           // ===============================================================
           // (7) SCAN REFERENCE ACQUISITION — pág. 10
           // FÍSICO: KUKA carga PN/frame y se coloca en el punto de INICIO de
           // la trayectoria de referencia. Tu lógica pone AtRefScanStart=TRUE cuando
           // está en posición. El PLC solo arma scan_ref_start si además los
           // parámetros mínimos (id_scan, x_size, y_size) están válidos (p. 10).
           // ===============================================================
       #cSTEP_SCAN_REF:

           // Validación mínima de parámetros de scan que el PLC publica al Supervisor
           #validScanParams := (LEN("PlcStatus".idScan) > 0) AND ("PlcStatus".xSize > 0.0) AND ("PlcStatus".ySize > 0.0);

           // Posicionar al inicio de Ref si no estamos (CASE 420, ARG=RefProgIdx)
           IF (NOT #kukaAtRefScanStartPos) AND (#WantCode_uint = 0) THEN
               #SupervisorCmdSeq := #SupervisorCmdSeq + 1;
               #WantCode_uint := #cKUKA_GOTO_REF_START; // ← KRC: CASE 420
               #WantProgRequestId := (#RefProgIdx);   // índice de programa REF por pieza
           END_IF;

           // Permiso de arranque
           IF #kukaAtRefScanStartPos AND #validScanParams AND NOT "SupervisorCmd".scanRefRunning THEN
               "PlcStatus".scanRefStart := TRUE;   // ← Anunciar “ready” al Supervisor
           END_IF;

           // Cuando el Supervisor arranca por primera vez → ejecutar trayectoria (CASE 432)
           IF (NOT #scanRefWasRunning) AND "SupervisorCmd".scanRefRunning THEN
               #SupervisorCmdSeq := #SupervisorCmdSeq + 1;
               #WantCode_uint := #cKUKA_RUN_REF_PATH;
               #WantProgRequestId := (#RefProgIdx);
           END_IF;

           IF "SupervisorCmd".scanRefRunning THEN
               #scanRefWasRunning := TRUE;
               IF #kukaRefScanFinished THEN
                   "PlcStatus".scanRefStart := FALSE;
               END_IF;
           END_IF;

           IF (NOT "SupervisorCmd".scanRefRunning) AND #scanRefWasRunning THEN
               #scanRefWasRunning := FALSE;
               "PlcStatus".scanRefStart := FALSE;

               IF NOT "SupervisorCmd".scanRefState THEN
                   "PlcStatus".stepPlc := #cSTEP_ID;
               ELSE
                   "PlcStatus".stepPlc := #cSTEP_SCAN_INSP;
               END_IF;
           END_IF;

           // ===============================================================
           // (8) SCAN INSPECTION — pág. 11
           // FÍSICO: KUKA se coloca en INICIO de la(s) trayectoria(s) de inspección
           // (AtInspScanStart=TRUE). El PLC arma scan_insp_start solo si parámetros
           // válidos. Supervisor corre/guarda y luego pide verificación (req_verif) (p. 11).
           // ===============================================================
       #cSTEP_SCAN_INSP:

           #validScanParams := (LEN("PlcStatus".idScan) > 0) AND ("PlcStatus".xSize > 0.0) AND ("PlcStatus".ySize > 0.0);

           // Posicionar al inicio de Insp (CASE 421, ARG=PartProgIdx)
           IF (NOT #kukaAtInspScanStartPos) AND (#WantCode_uint = 0) THEN
               #SupervisorCmdSeq := #SupervisorCmdSeq + 1;
               #WantCode_uint := #cKUKA_GOTO_INSP_START;
               #WantProgRequestId := (#PartProgIdx);
           END_IF;

           // Permiso de arranque
           IF #kukaAtInspScanStartPos AND #validScanParams AND NOT "SupervisorCmd".scanInsprunning THEN
               "PlcStatus".scanInspStart := TRUE;
           END_IF;

           // Al arrancar por primera vez → ejecutar trayectoria (CASE 433)
           IF (NOT #scanInspWasRunning) AND "SupervisorCmd".scanInsprunning THEN
               #SupervisorCmdSeq := #SupervisorCmdSeq + 1;
               #WantCode_uint := #cKUKA_RUN_INSP_PATH;
               #WantProgRequestId := (#PartProgIdx);
           END_IF;

           IF "SupervisorCmd".scanInsprunning THEN
               #scanInspWasRunning := TRUE;
               IF #kukaInspScanFinished THEN
                   "PlcStatus".scanInspStart := FALSE;
               END_IF;
           END_IF;

           IF (NOT "SupervisorCmd".scanInsprunning) AND #scanInspWasRunning THEN
               #scanInspWasRunning := FALSE;
               "PlcStatus".scanInspStart := FALSE;

               IF NOT "SupervisorCmd".scanInspState THEN
                   "PlcStatus".stepPlc := #cSTEP_ID;
               ELSE
                   // Pasar a verificación (latch)
                   IF "SupervisorCmd".reqVerif AND NOT #L_reqVerif THEN
                       "PlcStatus".stepPlc := #cSTEP_SCAN_REF_VERIF;
                       #L_reqVerif := TRUE;
                   END_IF;
                   IF NOT "SupervisorCmd".reqVerif THEN
                       #L_reqVerif := FALSE;
                   END_IF;
               END_IF;
           END_IF;


           // ===============================================================
           // (9) SCAN REFERENCE VERIFICATION — pág. 12
           // FÍSICO: KUKA vuelve al INICIO de la trayectoria de verificación de ref.
           // (AtRefScanStart=TRUE). Igual patrón de parámetros/ready/running/state (p. 12).
           // Fin: Supervisor decide Pre‑eval (req_pre_eval) o nuevo ciclo (req_identification_state).
           // ===============================================================
       #cSTEP_SCAN_REF_VERIF:

           #validScanParams := (LEN("PlcStatus".idScan) > 0) AND ("PlcStatus".xSize > 0.0) AND ("PlcStatus".ySize > 0.0);

           // Asegurar estar en inicio de Ref (CASE 420) antes de verificar
           IF (NOT #kukaAtRefScanStartPos) AND (#WantCode_uint = 0) THEN
               #SupervisorCmdSeq := #SupervisorCmdSeq + 1;
               #WantCode_uint := #cKUKA_GOTO_REF_START;
               #WantProgRequestId := (#RefProgIdx);
           END_IF;

           IF #kukaAtRefScanStartPos AND #validScanParams AND NOT "SupervisorCmd".scanRefRunning THEN
               "PlcStatus".scanRefStart := TRUE;
           END_IF;

           IF "SupervisorCmd".scanRefRunning THEN
               #scanRefWasRunning := TRUE;
           END_IF;

           IF (NOT "SupervisorCmd".scanRefRunning) AND #scanRefWasRunning THEN
               #scanRefWasRunning := FALSE;
               "PlcStatus".scanRefStart := FALSE;

               IF NOT "SupervisorCmd".scanRefState THEN
                   "PlcStatus".stepPlc := #cSTEP_ID;
               ELSE
                   // a) Pre‑eval
                   IF "SupervisorCmd".reqPreEval AND NOT #L_reqPreEval THEN
                       "PlcStatus".stepPlc := #cSTEP_PRE_EVAL;
                       #L_reqPreEval := TRUE;
                   END_IF;
                   IF NOT "SupervisorCmd".reqPreEval THEN
                       #L_reqPreEval := FALSE;
                   END_IF;

                   // b) Nuevo ciclo
                   IF "SupervisorCmd".reqIdentificationState AND NOT #L_reqIdent THEN
                       "PlcStatus".stepPlc := #cSTEP_ID;
                       #L_reqIdent := TRUE;
                   END_IF;
                   IF NOT "SupervisorCmd".reqIdentificationState THEN
                       #L_reqIdent := FALSE;
                   END_IF;
               END_IF;
           END_IF;

           // ===============================================================
           // (10) PRE‑EVALUATION / MARKING — pág. 13
           // FÍSICO: si la herramienta de marcado no está montada, el KUKA cambia
           // en Staübli al stand de “marking” según requiera el proceso; tras estar
           // listo se puede marcar (Supervisor.req_mark). El resultado físico del
           // marcado tu lógica lo refleja en MarkingDone=TRUE/FALSE (p. 13).
           // También se puede arrancar un nuevo ciclo (req_identification_state).
           // ===============================================================
       #cSTEP_PRE_EVAL:

           // Volver a Identification (una sola vez)
           IF "SupervisorCmd".reqIdentificationState AND NOT #L_reqIdent THEN
               "PlcStatus".stepPlc := #cSTEP_ID;
               #L_reqIdent := TRUE;
           END_IF;
           IF NOT "SupervisorCmd".reqIdentificationState THEN
               #L_reqIdent := FALSE;
           END_IF;

           // Marcado: un ciclo de ejecución por petición
           IF "SupervisorCmd".reqMark AND NOT #L_reqMark THEN
               "PlcStatus".markState := FALSE;
               "PlcStatus".markRunning := TRUE;
               "PlcStatus".markState := #MarkingDone;   // resultado físico del efector
               "PlcStatus".markRunning := FALSE;
               #L_reqMark := TRUE;
           END_IF;
           IF NOT "SupervisorCmd".reqMark THEN
               #L_reqMark := FALSE;
           END_IF;
       ELSE
           "PlcStatus".stepPlc := #cSTEP_ID;


   END_CASE;


   // ---------------------------------------------------------------
   // [2] DESPACHO AL KUKA (toggle goTrigger cuando el canal esté libre)
   //     • Este bloque “consume” el slot WantCmd → publica parámetros
   //       en los registros PNIO (con SWAP) → toggle de goTrigger.
   //     • El robot deberá igualar rbDone := goTrigger al terminar.
   // ---------------------------------------------------------------

   CASE #state OF
       0: // IDLE -> GO == ACK

           // "cancelGo" := FALSE;

           IF (#SupervisorCmdSeq <> #lastSeq) THEN

               IF  "goTrigger" = "rbDone" THEN

                   #code_int := #WantCode_uint;  // “code_int” que viajará al KRC

                   IF #code_int = 201 THEN
                       // id de herramienta → WORD+SWAP
                       // #Cfg_EndEffector
                       #toolReqId := SWAP(INT_TO_WORD(#WantToolRequestId));

                   END_IF;

                   IF #code_int = 414 THEN  //GOTO_TCG
                       // id de herramienta → WORD+SWAP
                       "requestIndexKuka" := SWAP(UINT_TO_WORD(#WantIndex));

                   END_IF;

                   IF #code_int = 420 THEN // GOTO_REF_START
                       // id de herramienta → WORD+SWAP
                       "programReqId" := SWAP(UINT_TO_WORD(#WantProgRequestId));

                   END_IF;

                   IF #code_int = 432 THEN // RUN_REF_PATH
                       // id de herramienta → WORD+SWAP
                       "programReqId" := SWAP(UINT_TO_WORD(#WantProgRequestId));

                   END_IF;

                   IF #code_int = 421 THEN // GOTO_REF_START
                       // id de herramienta → WORD+SWAP
                       "programReqId" := SWAP(UINT_TO_WORD(#WantProgRequestId));

                   END_IF;

                   IF #code_int = 433 THEN // RUN_INSP_PATH

                       "programReqId" := SWAP(UINT_TO_WORD(#WantProgRequestId));

                   END_IF;

                   // 2) Publicar código de movimiento
                   #moveCodeKuka := SWAP(UINT_TO_WORD(#code_int));   // KRC leerá "MoveCode" = INT

                   // 3) Disparo del GO: toggle de goTrigger (rbDone ≠ goTrigger → pedido activo)
                   "goTrigger" := NOT "goTrigger";

                   #lastSeq := #SupervisorCmdSeq;          // <-- memoriza!
                   #state := 20;

               END_IF;
           END_IF;

       20: // BUSY

           //#code_int := #KukaControlCmdCode;

           // CANCEL pedido en BUSY → avisar al KRC y ACK de la ORDEN ACTIVA
           IF #code_int = 903 THEN
               "cancelGo" := TRUE;
           END_IF;

           // Fin normal (o tras el cancel, cuando KRC cierra el canal por nivel)

           IF ("rbDone" = "goTrigger") THEN
               // 4) Vaciar slot de pendiente
               #WantCode_uint := 0;
               #WantProgRequestId := 0;
               #WantToolRequestId := 0;
               #WantIndex := 0;
               #state := 0;                            // vuelve a IDLE
           END_IF;

   END_CASE;
END_REGION
END_FUNCTION_BLOCK

ORGANIZATION_BLOCK "Main"   // OB1, LAD, ProgramCycle
TITLE = "Main Program Sweep (Cycle)"
{ S7_Optimized_Access := 'TRUE' }
VERSION : 0.1
   VAR_INPUT
      Initial_Call : Bool;   // Initial call of this OB
      Remanence : Bool;   // =True, if remanent data are available
   END_VAR
   VAR_TEMP
      evtEnterSrv : Bool;   // // Eventos de modo service jog
      evtEnterAuto : Bool;   // // Eventos de modo auto
      muxSelStb : Bool;
      muxStartStb : Bool;
      muxPgno : Byte;
      u : UDInt;
   END_VAR
BEGIN

REGION Network 1 (SCL): // ====================== READ (%I) ======================
   // // —— Enlaza estos símbolos a tus %I en el árbol de dispositivos ——
   //   // EStop_DI, SafeDoor_DI, AirPressure_DI, WaterInsp_DI, WaterTank_DI, RobotReady_DI, ...
   "$MOVE_ENABLE" := TRUE;
   "$I_O_ACT" := TRUE;
   //"$IN_HOME"
   //"$EXT"
   "PlcStatus".systemArmed := FALSE;
   "PlcStatus".robotInAutExt := "$EXT";
   "PlcStatus".robotInHome := "$IN_HOME";
END_REGION

REGION Network 2
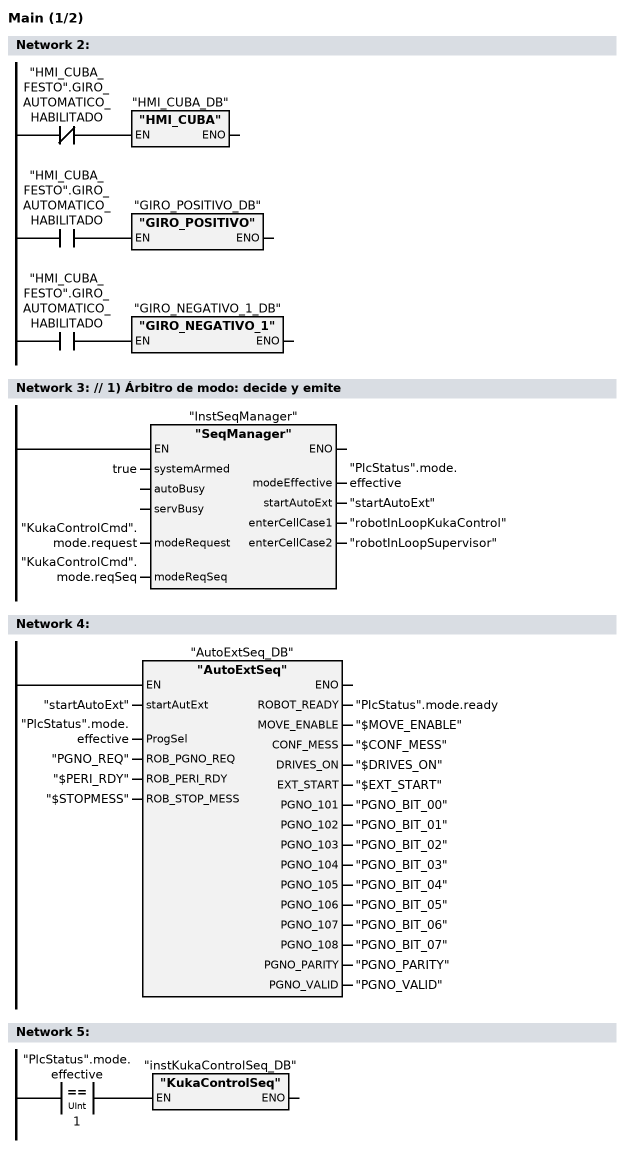
   RUNG wire#powerrail
      I_Contact( "HMI_CUBA_FESTO".GIRO_AUTOMATICO_HABILITADO )
      "HMI_CUBA_DB"()
   END_RUNG
   RUNG wire#powerrail
      Contact( "HMI_CUBA_FESTO".GIRO_AUTOMATICO_HABILITADO )
      "GIRO_POSITIVO_DB"()
   END_RUNG
   RUNG wire#powerrail
      Contact( "HMI_CUBA_FESTO".GIRO_AUTOMATICO_HABILITADO )
      "GIRO_NEGATIVO_1_DB"()
   END_RUNG
   // the same network as SCL:
   IF NOT "HMI_CUBA_FESTO".GIRO_AUTOMATICO_HABILITADO THEN
       "HMI_CUBA_DB"();   // "HMI_CUBA"
   END_IF;
   IF "HMI_CUBA_FESTO".GIRO_AUTOMATICO_HABILITADO THEN
       "GIRO_POSITIVO_DB"();   // "GIRO_POSITIVO"
   END_IF;
   IF "HMI_CUBA_FESTO".GIRO_AUTOMATICO_HABILITADO THEN
       "GIRO_NEGATIVO_1_DB"();   // "GIRO_NEGATIVO_1"
   END_IF;
END_REGION

REGION Network 3: // 1) Árbitro de modo: decide y emite
   RUNG wire#powerrail
      "InstSeqManager"(systemArmed := true, autoBusy :=, servBusy :=, modeRequest := "KukaControlCmd".mode.request, modeReqSeq := "KukaControlCmd".mode.reqSeq, modeEffective => "PlcStatus".mode.effective, startAutoExt => "startAutoExt", enterCellCase1 => "robotInLoopKukaControl", enterCellCase2 => "robotInLoopSupervisor")
   END_RUNG
   // the same network as SCL:
   "InstSeqManager"(systemArmed := true,   // "SeqManager"
                    modeRequest := "KukaControlCmd".mode.request,
                    modeReqSeq := "KukaControlCmd".mode.reqSeq,
                    modeEffective => "PlcStatus".mode.effective,
                    startAutoExt => "startAutoExt",
                    enterCellCase1 => "robotInLoopKukaControl",
                    enterCellCase2 => "robotInLoopSupervisor");
END_REGION

REGION Network 4
   RUNG wire#powerrail
      "AutoExtSeq_DB"(startAutExt := "startAutoExt", ProgSel := "PlcStatus".mode.effective, ROB_PGNO_REQ := "PGNO_REQ", ROB_PERI_RDY := "$PERI_RDY", ROB_STOP_MESS := "$STOPMESS", ROBOT_READY => "PlcStatus".mode.ready, MOVE_ENABLE => "$MOVE_ENABLE", CONF_MESS => "$CONF_MESS", DRIVES_ON => "$DRIVES_ON", EXT_START => "$EXT_START", PGNO_101 => "PGNO_BIT_00", PGNO_102 => "PGNO_BIT_01", PGNO_103 => "PGNO_BIT_02", PGNO_104 => "PGNO_BIT_03", PGNO_105 => "PGNO_BIT_04", PGNO_106 => "PGNO_BIT_05", PGNO_107 => "PGNO_BIT_06", PGNO_108 => "PGNO_BIT_07", PGNO_PARITY => "PGNO_PARITY", PGNO_VALID => "PGNO_VALID")
   END_RUNG
   // the same network as SCL:
   "AutoExtSeq_DB"(startAutExt := "startAutoExt",   // "AutoExtSeq"
                   ProgSel := "PlcStatus".mode.effective,
                   ROB_PGNO_REQ := "PGNO_REQ",
                   ROB_PERI_RDY := "$PERI_RDY",
                   ROB_STOP_MESS := "$STOPMESS",
                   ROBOT_READY => "PlcStatus".mode.ready,
                   MOVE_ENABLE => "$MOVE_ENABLE",
                   CONF_MESS => "$CONF_MESS",
                   DRIVES_ON => "$DRIVES_ON",
                   EXT_START => "$EXT_START",
                   PGNO_101 => "PGNO_BIT_00",
                   PGNO_102 => "PGNO_BIT_01",
                   PGNO_103 => "PGNO_BIT_02",
                   PGNO_104 => "PGNO_BIT_03",
                   PGNO_105 => "PGNO_BIT_04",
                   PGNO_106 => "PGNO_BIT_05",
                   PGNO_107 => "PGNO_BIT_06",
                   PGNO_108 => "PGNO_BIT_07",
                   PGNO_PARITY => "PGNO_PARITY",
                   PGNO_VALID => "PGNO_VALID");
END_REGION

REGION Network 5
   RUNG wire#powerrail
      { S7_Templates := "SrcType := UInt" } EQ_Contact(in1 := "PlcStatus".mode.effective, in2 := 1)
      "instKukaControlSeq_DB"()
   END_RUNG
   // the same network as SCL:
   IF "PlcStatus".mode.effective = 1 THEN
       "instKukaControlSeq_DB"();   // "KukaControlSeq"
   END_IF;
END_REGION

REGION Network 6
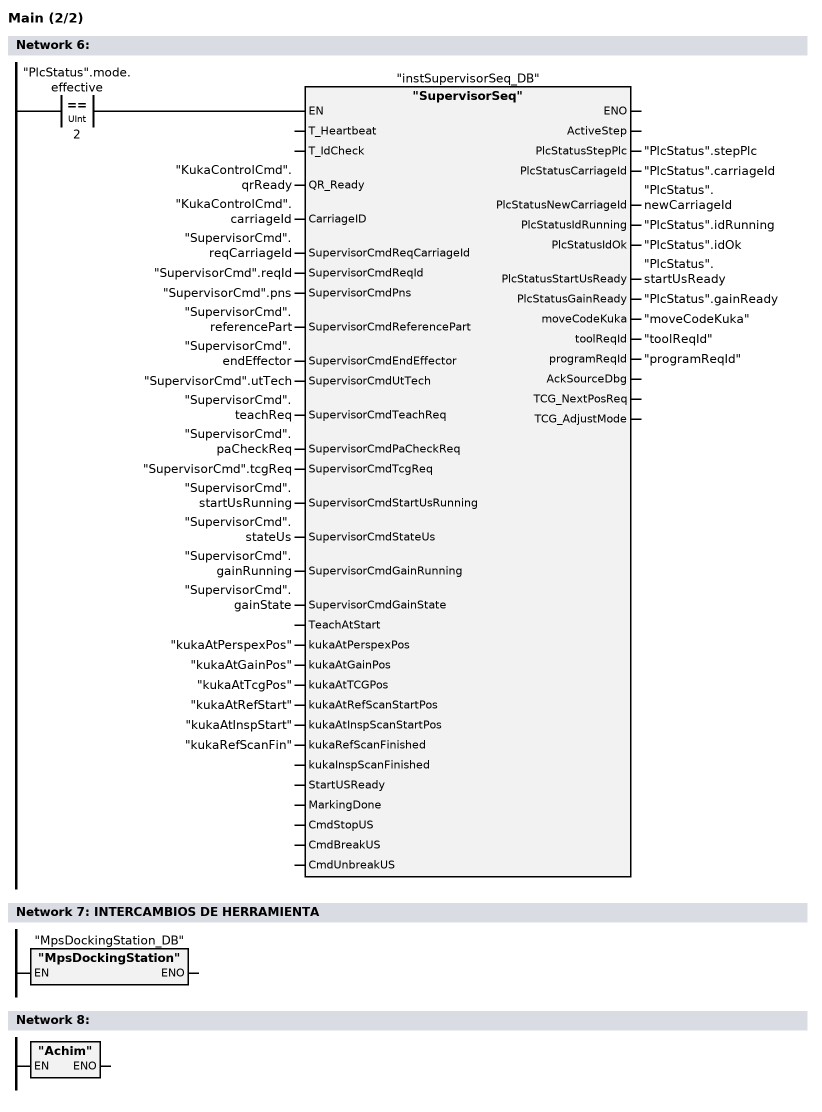
   RUNG wire#powerrail
      { S7_Templates := "SrcType := UInt" } EQ_Contact(in1 := "PlcStatus".mode.effective, in2 := 2)
      "instSupervisorSeq_DB"(T_Heartbeat :=, T_IdCheck :=, QR_Ready := "KukaControlCmd".qrReady, CarriageID := "KukaControlCmd".carriageId, SupervisorCmdReqCarriageId := "SupervisorCmd".reqCarriageId, SupervisorCmdReqId := "SupervisorCmd".reqId, SupervisorCmdPns := "SupervisorCmd".pns, SupervisorCmdReferencePart := "SupervisorCmd".referencePart, SupervisorCmdEndEffector := "SupervisorCmd".endEffector, SupervisorCmdUtTech := "SupervisorCmd".utTech, SupervisorCmdTeachReq := "SupervisorCmd".teachReq, SupervisorCmdPaCheckReq := "SupervisorCmd".paCheckReq, SupervisorCmdTcgReq := "SupervisorCmd".tcgReq, SupervisorCmdStartUsRunning := "SupervisorCmd".startUsRunning, SupervisorCmdStateUs := "SupervisorCmd".stateUs, SupervisorCmdGainRunning := "SupervisorCmd".gainRunning, SupervisorCmdGainState := "SupervisorCmd".gainState, TeachAtStart :=, kukaAtPerspexPos := "kukaAtPerspexPos", kukaAtGainPos := "kukaAtGainPos", kukaAtTCGPos := "kukaAtTcgPos", kukaAtRefScanStartPos := "kukaAtRefStart", kukaAtInspScanStartPos := "kukaAtInspStart", kukaRefScanFinished := "kukaRefScanFin", kukaInspScanFinished :=, StartUSReady :=, MarkingDone :=, CmdStopUS :=, CmdBreakUS :=, CmdUnbreakUS :=, ActiveStep =>, PlcStatusStepPlc => "PlcStatus".stepPlc, PlcStatusCarriageId => "PlcStatus".carriageId, PlcStatusNewCarriageId => "PlcStatus".newCarriageId, PlcStatusIdRunning => "PlcStatus".idRunning, PlcStatusIdOk => "PlcStatus".idOk, PlcStatusStartUsReady => "PlcStatus".startUsReady, PlcStatusGainReady => "PlcStatus".gainReady, moveCodeKuka => "moveCodeKuka", toolReqId => "toolReqId", programReqId => "programReqId", AckSourceDbg =>, TCG_NextPosReq =>, TCG_AdjustMode =>)
   END_RUNG
   // the same network as SCL:
   IF "PlcStatus".mode.effective = 2 THEN
       "instSupervisorSeq_DB"(QR_Ready := "KukaControlCmd".qrReady,   // "SupervisorSeq"
                              CarriageID := "KukaControlCmd".carriageId,
                              SupervisorCmdReqCarriageId := "SupervisorCmd".reqCarriageId,
                              SupervisorCmdReqId := "SupervisorCmd".reqId,
                              SupervisorCmdPns := "SupervisorCmd".pns,
                              SupervisorCmdReferencePart := "SupervisorCmd".referencePart,
                              SupervisorCmdEndEffector := "SupervisorCmd".endEffector,
                              SupervisorCmdUtTech := "SupervisorCmd".utTech,
                              SupervisorCmdTeachReq := "SupervisorCmd".teachReq,
                              SupervisorCmdPaCheckReq := "SupervisorCmd".paCheckReq,
                              SupervisorCmdTcgReq := "SupervisorCmd".tcgReq,
                              SupervisorCmdStartUsRunning := "SupervisorCmd".startUsRunning,
                              SupervisorCmdStateUs := "SupervisorCmd".stateUs,
                              SupervisorCmdGainRunning := "SupervisorCmd".gainRunning,
                              SupervisorCmdGainState := "SupervisorCmd".gainState,
                              kukaAtPerspexPos := "kukaAtPerspexPos",
                              kukaAtGainPos := "kukaAtGainPos",
                              kukaAtTCGPos := "kukaAtTcgPos",
                              kukaAtRefScanStartPos := "kukaAtRefStart",
                              kukaAtInspScanStartPos := "kukaAtInspStart",
                              kukaRefScanFinished := "kukaRefScanFin",
                              PlcStatusStepPlc => "PlcStatus".stepPlc,
                              PlcStatusCarriageId => "PlcStatus".carriageId,
                              PlcStatusNewCarriageId => "PlcStatus".newCarriageId,
                              PlcStatusIdRunning => "PlcStatus".idRunning,
                              PlcStatusIdOk => "PlcStatus".idOk,
                              PlcStatusStartUsReady => "PlcStatus".startUsReady,
                              PlcStatusGainReady => "PlcStatus".gainReady,
                              moveCodeKuka => "moveCodeKuka",
                              toolReqId => "toolReqId",
                              programReqId => "programReqId");
   END_IF;
END_REGION

REGION Network 7: INTERCAMBIOS DE HERRAMIENTA
   RUNG wire#powerrail
      "MpsDockingStation_DB"()
   END_RUNG
   // the same network as SCL:
   "MpsDockingStation_DB"();   // "MpsDockingStation"
END_REGION

REGION Network 8
   RUNG wire#powerrail
      "Achim"()
   END_RUNG
   // the same network as SCL:
   "Achim"();
END_REGION
END_ORGANIZATION_BLOCK

// folder: 20. Robot Services/AutoExt

FUNCTION_BLOCK "AutoExtSeq"   // FB31, LAD
{ S7_Optimized_Access := 'TRUE' }
VERSION : 0.1
   VAR_INPUT
      startAutExt : Bool;   // // Flanco para ejecutar CASE 1
      ProgSel : UInt;
      ROB_PGNO_REQ : Bool;
      ROB_PERI_RDY : Bool;
      ROB_STOP_MESS : Bool;
   END_VAR
   VAR_OUTPUT
      ROBOT_READY : Bool;
      MOVE_ENABLE : Bool := TRUE;
      CONF_MESS : Bool;
      DRIVES_ON : Bool;
      EXT_START : Bool;
      PGNO_101 : Bool;
      PGNO_102 : Bool;
      PGNO_103 : Bool;
      PGNO_104 : Bool;
      PGNO_105 : Bool;
      PGNO_106 : Bool;
      PGNO_107 : Bool;
      PGNO_108 : Bool;
      PGNO_PARITY : Bool;
      PGNO_VALID : Bool;
   END_VAR
   VAR
      "step" : Int;   // secuencia simple
      rStart : R_TRIG;
      rPgnoReq : R_TRIG;
      fPgnoReq : F_TRIG;
      tpConf : TP_TIME;
      tpDrives : TP_TIME;
      tpStart : TP_TIME;
      tpStartInit : TP_TIME;
      tStable : TON_TIME;
      pulseTime : Time := T#120ms;
      drivesPulse : Time := T#120ms;
      stableTime : Time := T#36ms;
      initStartPulse : Time := T#150ms;
      pgnoLatched : UInt;
      tPump : TP_TIME;
   END_VAR
BEGIN

REGION Network 1 (SCL): // === Secuencia Aut Ext ===
   /// 1) Detectores de flanco: se ejecutan SIEMPRE (cada ciclo de scan del plc)
   #rStart(CLK := #startAutExt);       // flanco de arranque de la secuencia
   #rPgnoReq(CLK := #ROB_PGNO_REQ);    // flanco de subida del PGNO_REQ
   #fPgnoReq(CLK := #ROB_PGNO_REQ);     // flanco de bajada del PGNO_REQ

   // 2) Valores por defecto de salidas “pulsadas” (evita retenerlas fuera de sus pasos)
   #DRIVES_ON := FALSE;
   #CONF_MESS := FALSE;
   #EXT_START := FALSE;


   // ------------------------------ Máquina de estados ---------------------
   CASE #step OF

       0:   // IDLE: esperar flanco de arranque externo (#startAutExt 0→1)

           // No imprescindible, pero dejamos los temporizadores “quietos”
           #tpStartInit(IN := FALSE,
                        PT := #initStartPulse);
           #tpDrives(IN := FALSE,
                     PT := #initStartPulse);
           #tpStart(IN := FALSE,
                    PT := #initStartPulse);

           // Por defecto, PGNO inválido en reposo  para iniciar “limpio”
           #PGNO_VALID := FALSE;

           // Poner a '0' los bits PGNO mientras no haya petición del KRC
           #PGNO_101 := FALSE;
           #PGNO_102 := FALSE;
           #PGNO_103 := FALSE;
           #PGNO_104 := FALSE;
           #PGNO_105 := FALSE;
           #PGNO_106 := FALSE;
           #PGNO_107 := FALSE;
           #PGNO_108 := FALSE;
           #PGNO_PARITY := FALSE;

           // Arrancar SOLO en flanco de #startAutExt
           IF #rStart.Q THEN // SOLO en el flanco  (un ciclo)
               #ROBOT_READY := FALSE;   // el modo no está listo mientras arranca
               #step := 1;               // → primer pulso: DRIVES_ON
           END_IF;


       1:  // Pulso de DRIVES_ON (una sola vez por ciclo de autoext)
           // Llamamos al TP solo en este paso ⇒ genera un único pulso de ancho #drivesPulse
           #tpDrives(IN := TRUE,
                     PT := #drivesPulse);
           #DRIVES_ON := #tpDrives.Q;
           IF NOT #tpDrives.Q THEN
               #step := 2;          // cuando cae el pulso → segundo pulso
           END_IF;


       2:  // Pulso de CONF_MESS (también una sola vez)
           #tpConf(IN := TRUE,
                   PT := #drivesPulse);   // o #confPulse si quieres ancho distinto
           #CONF_MESS := #tpConf.Q;
           IF NOT #tpConf.Q THEN
               #step := 5;           // luego hacemos el pre‑start (salir de INIT)
           END_IF;


       5:  // PRE‑START: salir de AUTOEXT INIT con un start corto
           #tpStartInit(IN := TRUE,
                        PT := #initStartPulse);
           #EXT_START := #tpStartInit.Q;
           IF NOT #tpStartInit.Q THEN
               #step := 10; // → esperar petición de PGNO por parte del KRC
           END_IF;

           // -------------------------------------------------------
       10: // Esperar a que el KRC pida número de programa (PGNO_REQ = 1)
           IF #ROB_PGNO_REQ THEN
               // Latch del programa seleccionado (1..3). Forzamos límites por seguridad.
               IF #ProgSel < USINT#1 THEN
                   #pgnoLatched := USINT#1;
               ELSIF #ProgSel > USINT#3 THEN
                   #pgnoLatched := USINT#3;
               ELSE
                   #pgnoLatched := #ProgSel;
               END_IF;

               #step := 20;
           END_IF;


       20: // Presentar PGNO MIENTRAS PGNO_REQ = 1
           IF #ROB_PGNO_REQ THEN
               // Escribir bits binarios 101..108 a partir de #pgnoLatched
               #PGNO_101 := ((#pgnoLatched AND USINT#1) <> USINT#0);
               #PGNO_102 := ((#pgnoLatched AND USINT#2) <> USINT#0);
               #PGNO_103 := ((#pgnoLatched AND USINT#4) <> USINT#0);
               #PGNO_104 := ((#pgnoLatched AND USINT#8) <> USINT#0);
               #PGNO_105 := ((#pgnoLatched AND USINT#16) <> USINT#0);
               #PGNO_106 := ((#pgnoLatched AND USINT#32) <> USINT#0);
               #PGNO_107 := ((#pgnoLatched AND USINT#64) <> USINT#0);
               #PGNO_108 := ((#pgnoLatched AND USINT#128) <> USINT#0);

               // Paridad "even": XOR de los 8 bits (1 si nº de unos es impar)
               #PGNO_PARITY :=
               #PGNO_101 XOR #PGNO_102 XOR #PGNO_103 XOR #PGNO_104 XOR
               #PGNO_105 XOR #PGNO_106 XOR #PGNO_107 XOR #PGNO_108;

               // Arrancamos el TON de estabilidad y pasamos a validación
               #tStable(IN := TRUE,
                        PT := #stableTime);
               #step := 21;
           END_IF;


       21: // Esperar estabilidad y marcar PGNO_VALID
           #tStable(IN := (#step = 21),
                    PT := #stableTime);
           IF #tStable.Q THEN
               #PGNO_VALID := TRUE;        // el KRC ya puede muestrear PGNO
               #step := 22;
           END_IF;


       22: // Mantener PGNO_VALID hasta la CAÍDA de PGNO_REQ
           #PGNO_VALID := TRUE;
           IF #fPgnoReq.Q THEN
               #PGNO_VALID := FALSE;    // cerrar handshake de selección

               // limpiar PGNO para siguientes ciclos
               #PGNO_101 := FALSE;
               #PGNO_102 := FALSE;
               #PGNO_103 := FALSE;
               #PGNO_104 := FALSE;
               #PGNO_105 := FALSE;
               #PGNO_106 := FALSE;
               #PGNO_107 := FALSE;
               #PGNO_108 := FALSE;
               #PGNO_PARITY := FALSE;

               #step := 40;    // → arranque real del programa
           END_IF;

       40: // START real: segundo pulso de $EXT_START para ejecutar el programa
           "Tag_10" := TRUE; // marcador/diagnóstico ELIMINAR
           #tpStart(IN := TRUE,
                    PT := #pulseTime);
           #EXT_START := #tpStart.Q;
           IF NOT #tpStart.Q THEN
               #ROBOT_READY := TRUE;   // handshake completo
               #step := 60;            // → ejecución
           END_IF;


       60: // En ejecución / rearme
           // Para un nuevo ciclo hay que hacer hacer 0→1 de nuevo desde la aplicacion 
           // si #startAutExt no baja, #rStart.Q no volverá a disparar.
           #step := 0;

   END_CASE;
END_REGION
END_FUNCTION_BLOCK

// folder: 20. Robot Services/Mov Manual

FUNCTION_BLOCK "TcpJogging"   // FB5, LAD
{ S7_Optimized_Access := 'TRUE' }
VERSION : 0.1
   VAR_INPUT
      "buttonX+" : Bool;
      "buttonX-" : Bool;
      "buttonY+" : Bool;
      "buttonY-" : Bool;
      "buttonZ+" : Bool;
      "buttonZ-" : Bool;
      "buttonE1+" : Bool;
      "buttonE1-" : Bool;
   END_VAR
BEGIN

REGION Network 1 (SCL): Mapea los valores de los botones de WF
   IF "PlcStatus".mode.effective = 0 THEN

       "Tag_1" := TRUE;
       //MOV X,Y,Z
       //%Q630.0 = buttonX+
       //%Q630.1 = buttonX-
       //%Q630.2 = buttonY+
       //%Q630.3 = buttonY-
       //%Q630.4 = buttonZ+
       //%Q630.5 = buttonZ-
       //MOV A,B,C
       //%Q630.6 = buttonWF +A
       //%Q630.7 = buttonWF -A
       //%Q631.0 = buttonWF +B
       //%Q631.1 = buttonWF -B
       //%Q631.2 = buttonWF +C
       //%Q631.3 = buttonWF -C
       //Mov E1
       //%Q631.4 = buttonWF +E1
       //%Q631.5 = buttonWF -E1

   ELSE
       //%Q631.1 = buttonWF -B
       "Tag_1" := FALSE;
   END_IF;
END_REGION
END_FUNCTION_BLOCK

FUNCTION_BLOCK "TcpTarget"   // FB11, LAD
{ S7_Optimized_Access := 'TRUE' }
VERSION : 0.1
   VAR_INPUT
      KukaControlCmdCode : UInt;
      KukaControlCmdSeq : UInt;
      KukaControlCmdProfileRequestId : UInt;
      KukaControlCmdToolRequestId : UInt;
      KukaControlCmdBaseRequestId : UInt;
      KukaControlCmdProgramRequestId : UInt;
      KukaControlTcpTargetX_mm : LReal;
      KukaControlTcpTargetY_mm : LReal;
      KukaControlTcpTargetZ_mm : LReal;
      kukaControlE1Target_mm : LReal;
      KukaControlCmdCancelGo : Bool;
      KukaControlCmdPauseGo : Bool;
      KukaControlCmdResumeGo : Bool;
      enterService : Bool;
      KukaControlCmdVel : UInt;
      KukaControlCmdIndex : UInt;
      scanPuntoInicialX : LReal;
      scanPuntoInicialY : LReal;
      scanPuntoInicialZ : LReal;
      scanPuntoInicialE1 : LReal;
      scanPuntoFinalX : LReal;
      scanPuntoFinalY : LReal;
      scanPuntoFinalZ : LReal;
      scanPuntoFinalE1 : LReal;
   END_VAR
   VAR_OUTPUT
      moveCodeKuka : Word;
      profileReqId : Word;
      baseReqId : Word;
      toolReqId : Word;
      programReqId : Word;
      x_mmHe : DWord;
      y_mmHe : DWord;
      z_mmHe : DWord;
      e_mmHe : DWord;
      PlcStatusExecDone : Bool;
      PlcStatusExecAccepted : Bool;
      PlcStatusExecAckSeq : UInt;
      PlcStatusExecBusy : Bool;
      PlcStatusExecError : Bool;
      PlcStatusExecErrorCode : DWord;
      PlcStatusExecLastCode : UInt;
      vel_mmsHe : Word;
      index_mmHe : Word;
      xInicial_mm : DWord;
      yInicial_mm : DWord;
      zInicial_mm : DWord;
      e1Inicial_mm : DWord;
      xFinal_mm : DWord;
      yFinal_mm : DWord;
      zFinal_mm : DWord;
      e1Final_mm : DWord;
   END_VAR
   VAR
      lastSeq : UInt;
      lastCode : UInt;
      state : Int;
      tmoMove : TON_TIME;
      rbDoneEdge : R_TRIG;
      _cancelInFlight : Bool := false;   // marca que el DONE que venga es por cancelación
      _isMotion : Bool;   // helper para saber si el code es de movimiento
      rbDoneEdge_1 : R_TRIG;
      rEnterSrv : R_TRIG;
   END_VAR
   VAR_TEMP
      x_dint : DInt;
      y_dint : DInt;
      z_dint : DInt;
      n_dint : DInt;
      code_int : UInt;
      tool_int : UInt;
      xInicial_dint : DInt;
      yInicial_Dint : DInt;
      ZInicial_Dint : DInt;
      e1Inicial_Dint : DInt;
      xFinal_Dint : DInt;
      yFinal_Dint : DInt;
      ZFinal_Dint : DInt;
      e1Final_Dint : DInt;
      index_uint : UInt;
      vel_uint : UInt;
   END_VAR
BEGIN

REGION Network 1 (SCL)
   #rEnterSrv(CLK := #enterService);
   IF #rEnterSrv.Q THEN
       #state := 0;
       #PlcStatusExecAccepted := FALSE;
       #PlcStatusExecBusy := FALSE;
       #PlcStatusExecDone := FALSE;

       // deja lastSeq "uno por detrás" del actual
       IF #KukaControlCmdSeq = UINT#0 THEN
           #lastSeq := UINT#65535;
       ELSE
           #lastSeq := #KukaControlCmdSeq - UINT#1;
       END_IF;
   END_IF;




   CASE #state OF
       0: // IDLE -> GO == ACK
           #PlcStatusExecAccepted := FALSE;
           #PlcStatusExecBusy := FALSE;
           #PlcStatusExecError := FALSE;
           "cancelGo" := FALSE;
           //#PlcStatusExecDone := FALSE;

           #code_int := #KukaControlCmdCode;  // refresca SIEMPRE

           #tool_int := #KukaControlCmdToolRequestId;

           // Nuevo comando si llega seq distinto y el canal está libre
           IF (#KukaControlCmdSeq <> #lastSeq) AND ("goTrigger" = "rbDone") THEN

                   IF #code_int = 130 THEN
                       //  Primero: Escalar mm → entero (µm). Ajusta el redondeo si lo prefieres TRUNC, FLOOR, etc.
                       #n_dint := LREAL_TO_DINT(ROUND(#kukaControlE1Target_mm));
                       // Segundo Convertir a DWORD y hacer SWAP para que el KRC lo lea correctamente
                       #e_mmHe := SWAP(DINT_TO_DWORD(#n_dint));
                   END_IF;

                   IF #code_int = 101 THEN
                       //  Primero: Escalar mm → entero (µm). Ajusta el redondeo si lo prefieres TRUNC, FLOOR, etc.
                       #x_dint := LREAL_TO_DINT(ROUND(#KukaControlTcpTargetX_mm));
                       // Segundo Convertir a DWORD y hacer SWAP para que el KRC lo lea correctamente
                       #x_mmHe := SWAP(DINT_TO_DWORD(#x_dint));
                   END_IF;

                   IF #code_int = 102 THEN
                       //  Primero: Escalar mm → entero (µm). Ajusta el redondeo si lo prefieres TRUNC, FLOOR, etc.
                       #y_dint := LREAL_TO_DINT(ROUND(#KukaControlTcpTargetY_mm));
                       // Segundo Convertir a DWORD y hacer SWAP para que el KRC lo lea correctamente
                       #y_mmHe := SWAP(DINT_TO_DWORD(#y_dint));
                   END_IF;

                   IF #code_int = 103 THEN
                       //  Primero: Escalar mm → entero (µm). Ajusta el redondeo si lo prefieres TRUNC, FLOOR, etc.
                       #z_dint := LREAL_TO_DINT(ROUND(#KukaControlTcpTargetZ_mm));
                       // Segundo Convertir a DWORD y hacer SWAP para que el KRC lo lea correctamente
                       #z_mmHe := SWAP(DINT_TO_DWORD(#z_dint));
                   END_IF;

                   IF #code_int = 201 THEN
                       // id de herramienta → WORD+SWAP
                       #toolReqId := SWAP(UINT_TO_WORD(#KukaControlCmdToolRequestId));

                   END_IF;

                   IF #code_int = 202 THEN

                       // id de herramienta → WORD+SWAP
                       #baseReqId := SWAP(UINT_TO_WORD(#KukaControlCmdBaseRequestId));

                   END_IF;

                   IF #code_int = 203 THEN

                       // id de herramienta → WORD+SWAP
                       #profileReqId := SWAP(UINT_TO_WORD(#KukaControlCmdProfileRequestId));

                   END_IF;

                   // ---------- TEACHING ----------
                   IF #code_int = 301 THEN // Teach Request
                       #programReqId := SWAP(UINT_TO_WORD(#KukaControlCmdProgramRequestId));

                   END_IF;

                   // ---------- TEACH SET START (desde SCA vía OPC) ----------
                   IF #code_int = 311 THEN

                       // Program ID (WORD + SWAP)
                       #programReqId := SWAP(UINT_TO_WORD(#KukaControlCmdProgramRequestId));


                       // Start desde OPC (mm -> DINT -> DWORD + SWAP)
                       //  Primero: Escalar mm → entero (µm). 
                       #xInicial_dint := LREAL_TO_DINT(ROUND(#scanPuntoInicialX));
                       // Segundo Convertir a DWORD y hacer SWAP para que el KRC lo lea correctamente
                       #xInicial_mm := SWAP(DINT_TO_DWORD(#xInicial_dint));
                       #yInicial_Dint := LREAL_TO_DINT(ROUND(#scanPuntoInicialY));
                       #yInicial_mm := SWAP(DINT_TO_DWORD(#yInicial_Dint));
                       #ZInicial_Dint := LREAL_TO_DINT(ROUND(#scanPuntoInicialZ));
                       #zInicial_mm := SWAP(DINT_TO_DWORD(#ZInicial_Dint));
                       #e1Inicial_Dint := LREAL_TO_DINT(ROUND(#scanPuntoInicialE1));
                       #e1Inicial_mm := SWAP(DINT_TO_DWORD(#e1Inicial_Dint));

                   END_IF;

                   // ---------- TEACH SET END (desde SCA vía OPC) ----------
                   IF #code_int = 312 THEN
                       // Program ID también aquí (por robustez)
                       #programReqId := SWAP(UINT_TO_WORD(#KukaControlCmdProgramRequestId));

                       // End desde OPC (mm -> DINT -> DWORD + SWAP)
                       #xFinal_Dint := LREAL_TO_DINT(ROUND(#scanPuntoFinalX));
                       #xFinal_mm := SWAP(DINT_TO_DWORD(#xFinal_Dint));
                       #yFinal_Dint := LREAL_TO_DINT(ROUND(#scanPuntoFinalY));
                       #yFinal_mm := SWAP(DINT_TO_DWORD(#yFinal_Dint));
                       #ZFinal_Dint := LREAL_TO_DINT(ROUND(#scanPuntoFinalZ));
                       #zFinal_mm := SWAP(DINT_TO_DWORD(#ZFinal_Dint));
                       #e1Final_Dint := LREAL_TO_DINT(ROUND(#scanPuntoFinalE1));
                       #e1Final_mm := SWAP(DINT_TO_DWORD(#e1Final_Dint));

                   END_IF;

                   // ---------- SCAN ----------
                   IF #code_int = 402 THEN

                       #programReqId := SWAP(UINT_TO_WORD(#KukaControlCmdProgramRequestId));

                       // ===== START: mm (LREAL) -> DINT -> DWORD + SWAP =====
                       #xInicial_dint := LREAL_TO_DINT(ROUND(#scanPuntoInicialX));
                       #xInicial_mm := SWAP(DINT_TO_DWORD(#xInicial_dint));

                       #yInicial_Dint := LREAL_TO_DINT(ROUND(#scanPuntoInicialY));
                       #yInicial_mm := SWAP(DINT_TO_DWORD(#yInicial_Dint));

                       #ZInicial_Dint := LREAL_TO_DINT(ROUND(#scanPuntoInicialZ));
                       #zInicial_mm := SWAP(DINT_TO_DWORD(#ZInicial_Dint));

                       #e1Inicial_Dint := LREAL_TO_DINT(ROUND(#scanPuntoInicialE1));
                       #e1Inicial_mm := SWAP(DINT_TO_DWORD(#e1Inicial_Dint));

                       // ===== END: mm (LREAL) -> DINT -> DWORD + SWAP =====
                       #xFinal_Dint := LREAL_TO_DINT(ROUND(#scanPuntoFinalX));
                       #xFinal_mm := SWAP(DINT_TO_DWORD(#xFinal_Dint));

                       #yFinal_Dint := LREAL_TO_DINT(ROUND(#scanPuntoFinalY));
                       #yFinal_mm := SWAP(DINT_TO_DWORD(#yFinal_Dint));

                       #ZFinal_Dint := LREAL_TO_DINT(ROUND(#scanPuntoFinalZ));
                       #zFinal_mm := SWAP(DINT_TO_DWORD(#ZFinal_Dint));

                       #e1Final_Dint := LREAL_TO_DINT(ROUND(#scanPuntoFinalE1));
                       #e1Final_mm := SWAP(DINT_TO_DWORD(#e1Final_Dint));

                       // ===== Opcional pero recomendado: velocidad e índice =====
                       // Si en KRC tienes mapeadas variables para vel/index:
                       #vel_uint := #KukaControlCmdVel;
                       #index_uint := #KukaControlCmdIndex;
                       #vel_mmsHe := SWAP(UINT_TO_WORD(#vel_uint));
                       #index_mmHe := SWAP(UINT_TO_WORD(#index_uint));
                       // #index_Dint  := LREAL_TO_DINT(ROUND(#KukaControlCmd_index_mm));
                       // #index_mmHe  := SWAP(DINT_TO_DWORD(#index_Dint));

                   END_IF;

